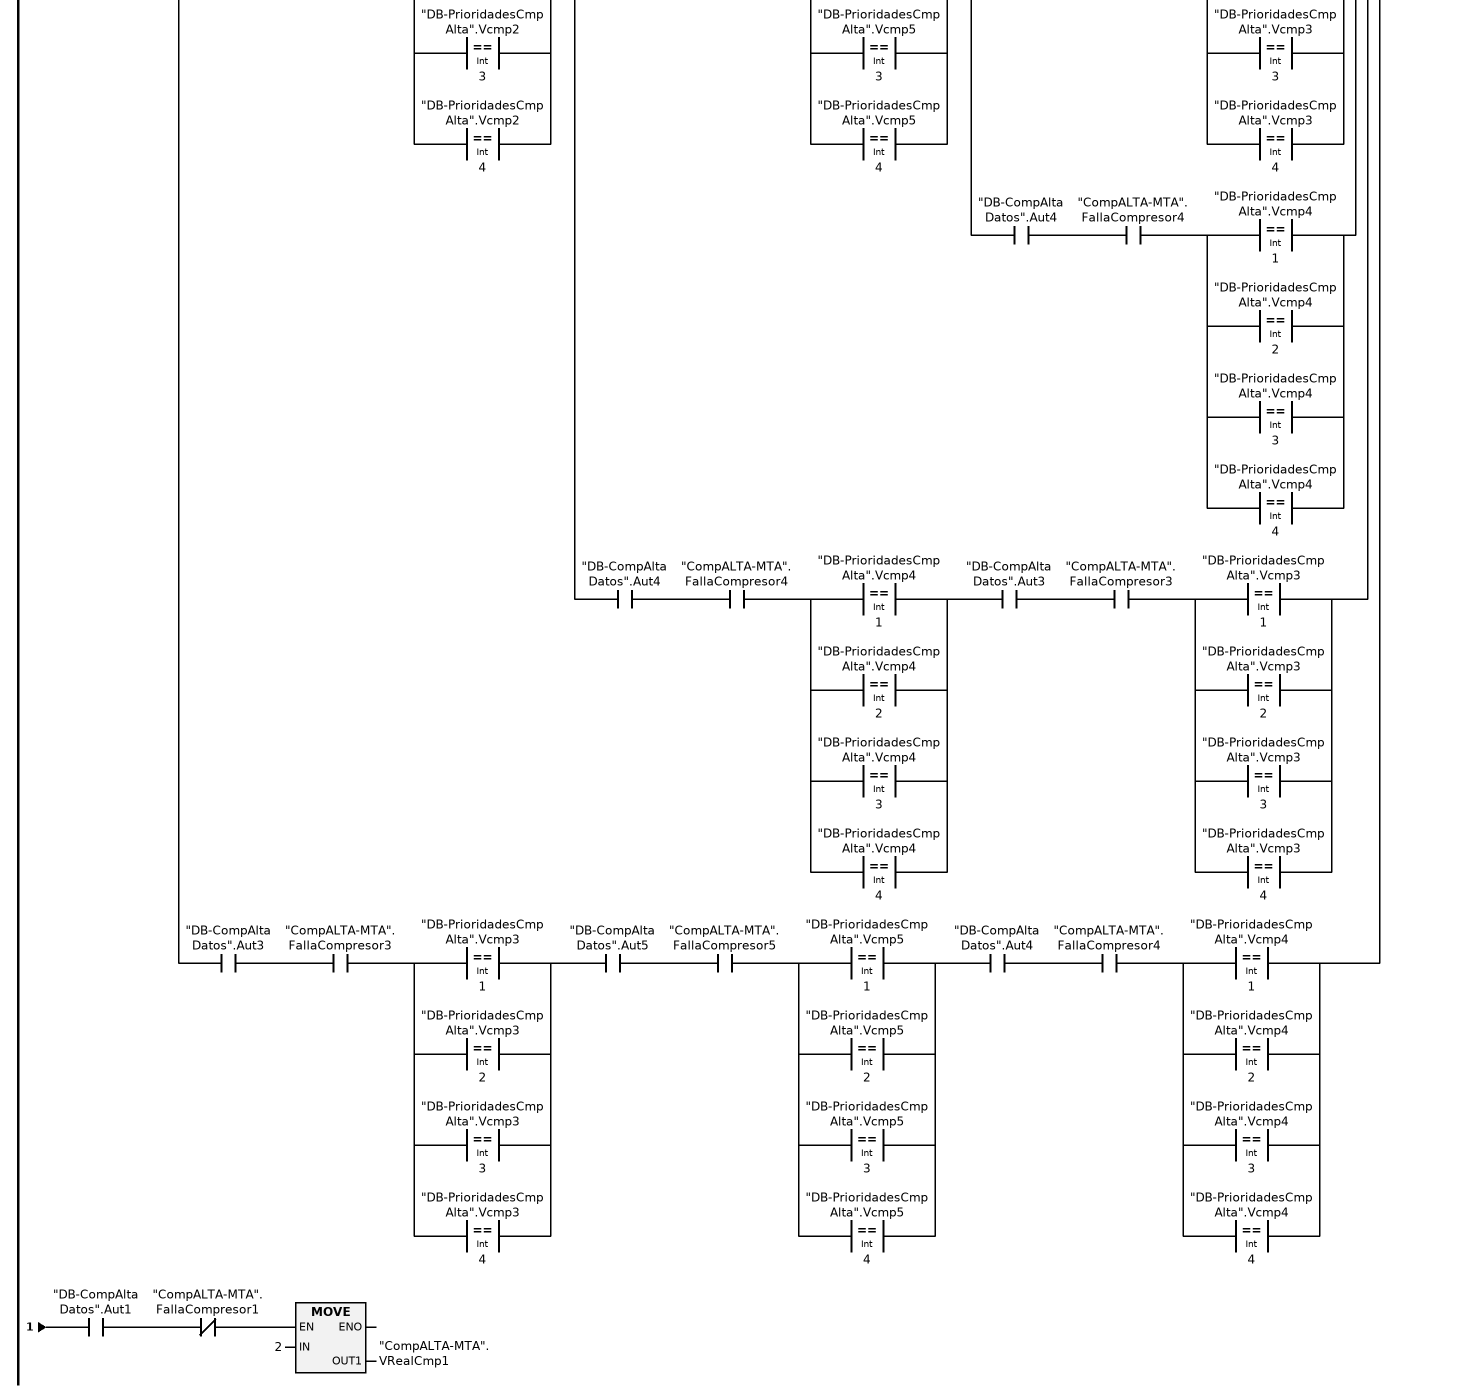
   RUNG wire#powerrail
      { S7_Templates := "SrcType := Int" } EQ_Contact(in1 := "DB-PrioridadesCmpAlta".Vcmp1, in2 := 2)
      wire#w1
      Contact( "DB-CompAltaDatos".Aut1 )
      I_Contact( "CompALTA-MTA".FallaCompresor1 )
      { S7_GenerateENO := "TRUE" } Move(in := 2, out1 => "CompALTA-MTA".VRealCmp1)
   END_RUNG
   RUNG wire#powerrail
      { S7_Templates := "SrcType := Int" } EQ_Contact(in1 := "DB-PrioridadesCmpAlta".Vcmp1, in2 := 3)
      wire#w2
      Contact( "DB-CompAltaDatos".Aut2 )
      Contact( "CompALTA-MTA".FallaCompresor2 )
      wire#w3
      { S7_Templates := "SrcType := Int" } EQ_Contact(in1 := "DB-PrioridadesCmpAlta".Vcmp2, in2 := 2)
   END_RUNG wire#w1
   RUNG wire#w3
      { S7_Templates := "SrcType := Int" } EQ_Contact(in1 := "DB-PrioridadesCmpAlta".Vcmp2, in2 := 1)
   END_RUNG wire#w1
   RUNG wire#w2
      Contact( "DB-CompAltaDatos".Aut3 )
      Contact( "CompALTA-MTA".FallaCompresor3 )
      wire#w4
      { S7_Templates := "SrcType := Int" } EQ_Contact(in1 := "DB-PrioridadesCmpAlta".Vcmp3, in2 := 2)
   END_RUNG wire#w1
   RUNG wire#w4
      { S7_Templates := "SrcType := Int" } EQ_Contact(in1 := "DB-PrioridadesCmpAlta".Vcmp3, in2 := 1)
   END_RUNG wire#w1
   RUNG wire#w2
      Contact( "DB-CompAltaDatos".Aut4 )
      Contact( "CompALTA-MTA".FallaCompresor4 )
      wire#w5
      { S7_Templates := "SrcType := Int" } EQ_Contact(in1 := "DB-PrioridadesCmpAlta".Vcmp4, in2 := 2)
   END_RUNG wire#w1
   RUNG wire#w5
      { S7_Templates := "SrcType := Int" } EQ_Contact(in1 := "DB-PrioridadesCmpAlta".Vcmp4, in2 := 1)
   END_RUNG wire#w1
   RUNG wire#w2
      Contact( "DB-CompAltaDatos".Aut5 )
      Contact( "CompALTA-MTA".FallaCompresor5 )
      wire#w6
      { S7_Templates := "SrcType := Int" } EQ_Contact(in1 := "DB-PrioridadesCmpAlta".Vcmp5, in2 := 2)
   END_RUNG wire#w1
   RUNG wire#w6
      { S7_Templates := "SrcType := Int" } EQ_Contact(in1 := "DB-PrioridadesCmpAlta".Vcmp5, in2 := 1)
   END_RUNG wire#w1
   RUNG wire#powerrail
      { S7_Templates := "SrcType := Int" } EQ_Contact(in1 := "DB-PrioridadesCmpAlta".Vcmp1, in2 := 4)
      wire#w7
      Contact( "DB-CompAltaDatos".Aut2 )
      Contact( "CompALTA-MTA".FallaCompresor2 )
      wire#w8
      { S7_Templates := "SrcType := Int" } EQ_Contact(in1 := "DB-PrioridadesCmpAlta".Vcmp2, in2 := 1)
      wire#w9
      Contact( "DB-CompAltaDatos".Aut5 )
      Contact( "CompALTA-MTA".FallaCompresor5 )
      wire#w10
      { S7_Templates := "SrcType := Int" } EQ_Contact(in1 := "DB-PrioridadesCmpAlta".Vcmp5, in2 := 1)
   END_RUNG wire#w1
   RUNG wire#w8
      { S7_Templates := "SrcType := Int" } EQ_Contact(in1 := "DB-PrioridadesCmpAlta".Vcmp2, in2 := 2)
   END_RUNG wire#w9
   RUNG wire#w8
      { S7_Templates := "SrcType := Int" } EQ_Contact(in1 := "DB-PrioridadesCmpAlta".Vcmp2, in2 := 3)
   END_RUNG wire#w9
   RUNG wire#w10
      { S7_Templates := "SrcType := Int" } EQ_Contact(in1 := "DB-PrioridadesCmpAlta".Vcmp5, in2 := 2)
   END_RUNG wire#w1
   RUNG wire#w10
      { S7_Templates := "SrcType := Int" } EQ_Contact(in1 := "DB-PrioridadesCmpAlta".Vcmp5, in2 := 3)
   END_RUNG wire#w1
   RUNG wire#w9
      Contact( "DB-CompAltaDatos".Aut4 )
      Contact( "CompALTA-MTA".FallaCompresor4 )
      wire#w11
      { S7_Templates := "SrcType := Int" } EQ_Contact(in1 := "DB-PrioridadesCmpAlta".Vcmp4, in2 := 1)
   END_RUNG wire#w1
   RUNG wire#w11
      { S7_Templates := "SrcType := Int" } EQ_Contact(in1 := "DB-PrioridadesCmpAlta".Vcmp4, in2 := 2)
   END_RUNG wire#w1
   RUNG wire#w11
      { S7_Templates := "SrcType := Int" } EQ_Contact(in1 := "DB-PrioridadesCmpAlta".Vcmp4, in2 := 3)
   END_RUNG wire#w1
   RUNG wire#w9
      Contact( "DB-CompAltaDatos".Aut3 )
      Contact( "CompALTA-MTA".FallaCompresor3 )
      wire#w12
      { S7_Templates := "SrcType := Int" } EQ_Contact(in1 := "DB-PrioridadesCmpAlta".Vcmp3, in2 := 1)
   END_RUNG wire#w1
   RUNG wire#w12
      { S7_Templates := "SrcType := Int" } EQ_Contact(in1 := "DB-PrioridadesCmpAlta".Vcmp3, in2 := 2)
   END_RUNG wire#w1
   RUNG wire#w12
      { S7_Templates := "SrcType := Int" } EQ_Contact(in1 := "DB-PrioridadesCmpAlta".Vcmp3, in2 := 3)
   END_RUNG wire#w1
   RUNG wire#w7
      Contact( "DB-CompAltaDatos".Aut3 )
      Contact( "CompALTA-MTA".FallaCompresor3 )
      wire#w13
      { S7_Templates := "SrcType := Int" } EQ_Contact(in1 := "DB-PrioridadesCmpAlta".Vcmp3, in2 := 1)
      wire#w14
      Contact( "DB-CompAltaDatos".Aut5 )
      Contact( "CompALTA-MTA".FallaCompresor5 )
      wire#w15
      { S7_Templates := "SrcType := Int" } EQ_Contact(in1 := "DB-PrioridadesCmpAlta".Vcmp5, in2 := 1)
   END_RUNG wire#w1
   RUNG wire#w13
      { S7_Templates := "SrcType := Int" } EQ_Contact(in1 := "DB-PrioridadesCmpAlta".Vcmp3, in2 := 2)
   END_RUNG wire#w14
   RUNG wire#w13
      { S7_Templates := "SrcType := Int" } EQ_Contact(in1 := "DB-PrioridadesCmpAlta".Vcmp3, in2 := 3)
   END_RUNG wire#w14
   RUNG wire#w15
      { S7_Templates := "SrcType := Int" } EQ_Contact(in1 := "DB-PrioridadesCmpAlta".Vcmp5, in2 := 2)
   END_RUNG wire#w1
   RUNG wire#w15
      { S7_Templates := "SrcType := Int" } EQ_Contact(in1 := "DB-PrioridadesCmpAlta".Vcmp5, in2 := 3)
   END_RUNG wire#w1
   RUNG wire#w14
      Contact( "DB-CompAltaDatos".Aut4 )
      Contact( "CompALTA-MTA".FallaCompresor4 )
      wire#w16
      { S7_Templates := "SrcType := Int" } EQ_Contact(in1 := "DB-PrioridadesCmpAlta".Vcmp4, in2 := 1)
   END_RUNG wire#w1
   RUNG wire#w16
      { S7_Templates := "SrcType := Int" } EQ_Contact(in1 := "DB-PrioridadesCmpAlta".Vcmp4, in2 := 2)
   END_RUNG wire#w1
   RUNG wire#w16
      { S7_Templates := "SrcType := Int" } EQ_Contact(in1 := "DB-PrioridadesCmpAlta".Vcmp4, in2 := 3)
   END_RUNG wire#w1
   RUNG wire#w7
      Contact( "DB-CompAltaDatos".Aut4 )
      Contact( "CompALTA-MTA".FallaCompresor4 )
      wire#w17
      { S7_Templates := "SrcType := Int" } EQ_Contact(in1 := "DB-PrioridadesCmpAlta".Vcmp4, in2 := 1)
      wire#w18
      Contact( "DB-CompAltaDatos".Aut5 )
      Contact( "CompALTA-MTA".FallaCompresor5 )
      wire#w19
      { S7_Templates := "SrcType := Int" } EQ_Contact(in1 := "DB-PrioridadesCmpAlta".Vcmp5, in2 := 1)
   END_RUNG wire#w1
   RUNG wire#w17
      { S7_Templates := "SrcType := Int" } EQ_Contact(in1 := "DB-PrioridadesCmpAlta".Vcmp4, in2 := 2)
   END_RUNG wire#w18
   RUNG wire#w17
      { S7_Templates := "SrcType := Int" } EQ_Contact(in1 := "DB-PrioridadesCmpAlta".Vcmp4, in2 := 3)
   END_RUNG wire#w18
   RUNG wire#w19
      { S7_Templates := "SrcType := Int" } EQ_Contact(in1 := "DB-PrioridadesCmpAlta".Vcmp5, in2 := 2)
   END_RUNG wire#w1
   RUNG wire#w19
      { S7_Templates := "SrcType := Int" } EQ_Contact(in1 := "DB-PrioridadesCmpAlta".Vcmp5, in2 := 3)
   END_RUNG wire#w1
   RUNG wire#powerrail
      { S7_Templates := "SrcType := Int" } EQ_Contact(in1 := "DB-PrioridadesCmpAlta".Vcmp1, in2 := 5)
      wire#w20
      Contact( "DB-CompAltaDatos".Aut2 )
      Contact( "CompALTA-MTA".FallaCompresor2 )
      wire#w21
      { S7_Templates := "SrcType := Int" } EQ_Contact(in1 := "DB-PrioridadesCmpAlta".Vcmp2, in2 := 1)
      wire#w22
      Contact( "DB-CompAltaDatos".Aut5 )
      Contact( "CompALTA-MTA".FallaCompresor5 )
      wire#w23
      { S7_Templates := "SrcType := Int" } EQ_Contact(in1 := "DB-PrioridadesCmpAlta".Vcmp5, in2 := 1)
      wire#w24
      Contact( "DB-CompAltaDatos".Aut3 )
      Contact( "CompALTA-MTA".FallaCompresor3 )
      wire#w25
      { S7_Templates := "SrcType := Int" } EQ_Contact(in1 := "DB-PrioridadesCmpAlta".Vcmp3, in2 := 1)
   END_RUNG wire#w1
   RUNG wire#w21
      { S7_Templates := "SrcType := Int" } EQ_Contact(in1 := "DB-PrioridadesCmpAlta".Vcmp2, in2 := 2)
   END_RUNG wire#w22
   RUNG wire#w21
      { S7_Templates := "SrcType := Int" } EQ_Contact(in1 := "DB-PrioridadesCmpAlta".Vcmp2, in2 := 3)
   END_RUNG wire#w22
   RUNG wire#w21
      { S7_Templates := "SrcType := Int" } EQ_Contact(in1 := "DB-PrioridadesCmpAlta".Vcmp2, in2 := 4)
   END_RUNG wire#w22
   RUNG wire#w23
      { S7_Templates := "SrcType := Int" } EQ_Contact(in1 := "DB-PrioridadesCmpAlta".Vcmp5, in2 := 2)
   END_RUNG wire#w24
   RUNG wire#w23
      { S7_Templates := "SrcType := Int" } EQ_Contact(in1 := "DB-PrioridadesCmpAlta".Vcmp5, in2 := 3)
   END_RUNG wire#w24
   RUNG wire#w23
      { S7_Templates := "SrcType := Int" } EQ_Contact(in1 := "DB-PrioridadesCmpAlta".Vcmp5, in2 := 4)
   END_RUNG wire#w24
   RUNG wire#w25
      { S7_Templates := "SrcType := Int" } EQ_Contact(in1 := "DB-PrioridadesCmpAlta".Vcmp3, in2 := 2)
   END_RUNG wire#w1
   RUNG wire#w25
      { S7_Templates := "SrcType := Int" } EQ_Contact(in1 := "DB-PrioridadesCmpAlta".Vcmp3, in2 := 3)
   END_RUNG wire#w1
   RUNG wire#w25
      { S7_Templates := "SrcType := Int" } EQ_Contact(in1 := "DB-PrioridadesCmpAlta".Vcmp3, in2 := 4)
   END_RUNG wire#w1
   RUNG wire#w24
      Contact( "DB-CompAltaDatos".Aut4 )
      Contact( "CompALTA-MTA".FallaCompresor4 )
      wire#w26
      { S7_Templates := "SrcType := Int" } EQ_Contact(in1 := "DB-PrioridadesCmpAlta".Vcmp4, in2 := 1)
   END_RUNG wire#w1
   RUNG wire#w26
      { S7_Templates := "SrcType := Int" } EQ_Contact(in1 := "DB-PrioridadesCmpAlta".Vcmp4, in2 := 2)
   END_RUNG wire#w1
   RUNG wire#w26
      { S7_Templates := "SrcType := Int" } EQ_Contact(in1 := "DB-PrioridadesCmpAlta".Vcmp4, in2 := 3)
   END_RUNG wire#w1
   RUNG wire#w26
      { S7_Templates := "SrcType := Int" } EQ_Contact(in1 := "DB-PrioridadesCmpAlta".Vcmp4, in2 := 4)
   END_RUNG wire#w1
   RUNG wire#w22
      Contact( "DB-CompAltaDatos".Aut4 )
      Contact( "CompALTA-MTA".FallaCompresor4 )
      wire#w27
      { S7_Templates := "SrcType := Int" } EQ_Contact(in1 := "DB-PrioridadesCmpAlta".Vcmp4, in2 := 1)
      wire#w28
      Contact( "DB-CompAltaDatos".Aut3 )
      Contact( "CompALTA-MTA".FallaCompresor3 )
      wire#w29
      { S7_Templates := "SrcType := Int" } EQ_Contact(in1 := "DB-PrioridadesCmpAlta".Vcmp3, in2 := 1)
   END_RUNG wire#w1
   RUNG wire#w27
      { S7_Templates := "SrcType := Int" } EQ_Contact(in1 := "DB-PrioridadesCmpAlta".Vcmp4, in2 := 2)
   END_RUNG wire#w28
   RUNG wire#w27
      { S7_Templates := "SrcType := Int" } EQ_Contact(in1 := "DB-PrioridadesCmpAlta".Vcmp4, in2 := 3)
   END_RUNG wire#w28
   RUNG wire#w27
      { S7_Templates := "SrcType := Int" } EQ_Contact(in1 := "DB-PrioridadesCmpAlta".Vcmp4, in2 := 4)
   END_RUNG wire#w28
   RUNG wire#w29
      { S7_Templates := "SrcType := Int" } EQ_Contact(in1 := "DB-PrioridadesCmpAlta".Vcmp3, in2 := 2)
   END_RUNG wire#w1
   RUNG wire#w29
      { S7_Templates := "SrcType := Int" } EQ_Contact(in1 := "DB-PrioridadesCmpAlta".Vcmp3, in2 := 3)
   END_RUNG wire#w1
   RUNG wire#w29
      { S7_Templates := "SrcType := Int" } EQ_Contact(in1 := "DB-PrioridadesCmpAlta".Vcmp3, in2 := 4)
   END_RUNG wire#w1
   RUNG wire#w20
      Contact( "DB-CompAltaDatos".Aut3 )
      Contact( "CompALTA-MTA".FallaCompresor3 )
      wire#w30
      { S7_Templates := "SrcType := Int" } EQ_Contact(in1 := "DB-PrioridadesCmpAlta".Vcmp3, in2 := 1)
      wire#w31
      Contact( "DB-CompAltaDatos".Aut5 )
      Contact( "CompALTA-MTA".FallaCompresor5 )
      wire#w32
      { S7_Templates := "SrcType := Int" } EQ_Contact(in1 := "DB-PrioridadesCmpAlta".Vcmp5, in2 := 1)
      wire#w33
      Contact( "DB-CompAltaDatos".Aut4 )
      Contact( "CompALTA-MTA".FallaCompresor4 )
      wire#w34
      { S7_Templates := "SrcType := Int" } EQ_Contact(in1 := "DB-PrioridadesCmpAlta".Vcmp4, in2 := 1)
   END_RUNG wire#w1
   RUNG wire#w30
      { S7_Templates := "SrcType := Int" } EQ_Contact(in1 := "DB-PrioridadesCmpAlta".Vcmp3, in2 := 2)
   END_RUNG wire#w31
   RUNG wire#w30
      { S7_Templates := "SrcType := Int" } EQ_Contact(in1 := "DB-PrioridadesCmpAlta".Vcmp3, in2 := 3)
   END_RUNG wire#w31
   RUNG wire#w30
      { S7_Templates := "SrcType := Int" } EQ_Contact(in1 := "DB-PrioridadesCmpAlta".Vcmp3, in2 := 4)
   END_RUNG wire#w31
   RUNG wire#w32
      { S7_Templates := "SrcType := Int" } EQ_Contact(in1 := "DB-PrioridadesCmpAlta".Vcmp5, in2 := 2)
   END_RUNG wire#w33
   RUNG wire#w32
      { S7_Templates := "SrcType := Int" } EQ_Contact(in1 := "DB-PrioridadesCmpAlta".Vcmp5, in2 := 3)
   END_RUNG wire#w33
   RUNG wire#w32
      { S7_Templates := "SrcType := Int" } EQ_Contact(in1 := "DB-PrioridadesCmpAlta".Vcmp5, in2 := 4)
   END_RUNG wire#w33
   RUNG wire#w34
      { S7_Templates := "SrcType := Int" } EQ_Contact(in1 := "DB-PrioridadesCmpAlta".Vcmp4, in2 := 2)
   END_RUNG wire#w1
   RUNG wire#w34
      { S7_Templates := "SrcType := Int" } EQ_Contact(in1 := "DB-PrioridadesCmpAlta".Vcmp4, in2 := 3)
   END_RUNG wire#w1
   RUNG wire#w34
      { S7_Templates := "SrcType := Int" } EQ_Contact(in1 := "DB-PrioridadesCmpAlta".Vcmp4, in2 := 4)
   END_RUNG wire#w1
   // the same network as SCL:
   IF (("DB-PrioridadesCmpAlta".Vcmp1 = 2) OR (("DB-PrioridadesCmpAlta".Vcmp1 = 3) AND (("DB-CompAltaDatos".Aut2 AND "CompALTA-MTA".FallaCompresor2 AND (("DB-PrioridadesCmpAlta".Vcmp2 = 2) OR ("DB-PrioridadesCmpAlta".Vcmp2 = 1))) OR ("DB-CompAltaDatos".Aut3 AND "CompALTA-MTA".FallaCompresor3 AND (("DB-PrioridadesCmpAlta".Vcmp3 = 2) OR ("DB-PrioridadesCmpAlta".Vcmp3 = 1))) OR ("DB-CompAltaDatos".Aut4 AND "CompALTA-MTA".FallaCompresor4 AND (("DB-PrioridadesCmpAlta".Vcmp4 = 2) OR ("DB-PrioridadesCmpAlta".Vcmp4 = 1))) OR ("DB-CompAltaDatos".Aut5 AND "CompALTA-MTA".FallaCompresor5 AND (("DB-PrioridadesCmpAlta".Vcmp5 = 2) OR ("DB-PrioridadesCmpAlta".Vcmp5 = 1))))) OR (("DB-PrioridadesCmpAlta".Vcmp1 = 4) AND (("DB-CompAltaDatos".Aut2 AND "CompALTA-MTA".FallaCompresor2 AND (("DB-PrioridadesCmpAlta".Vcmp2 = 1) OR ("DB-PrioridadesCmpAlta".Vcmp2 = 2) OR ("DB-PrioridadesCmpAlta".Vcmp2 = 3)) AND (("DB-CompAltaDatos".Aut5 AND "CompALTA-MTA".FallaCompresor5 AND (("DB-PrioridadesCmpAlta".Vcmp5 = 1) OR ("DB-PrioridadesCmpAlta".Vcmp5 = 2) OR ("DB-PrioridadesCmpAlta".Vcmp5 = 3))) OR ("DB-CompAltaDatos".Aut4 AND "CompALTA-MTA".FallaCompresor4 AND (("DB-PrioridadesCmpAlta".Vcmp4 = 1) OR ("DB-PrioridadesCmpAlta".Vcmp4 = 2) OR ("DB-PrioridadesCmpAlta".Vcmp4 = 3))) OR ("DB-CompAltaDatos".Aut3 AND "CompALTA-MTA".FallaCompresor3 AND (("DB-PrioridadesCmpAlta".Vcmp3 = 1) OR ("DB-PrioridadesCmpAlta".Vcmp3 = 2) OR ("DB-PrioridadesCmpAlta".Vcmp3 = 3))))) OR ("DB-CompAltaDatos".Aut3 AND "CompALTA-MTA".FallaCompresor3 AND (("DB-PrioridadesCmpAlta".Vcmp3 = 1) OR ("DB-PrioridadesCmpAlta".Vcmp3 = 2) OR ("DB-PrioridadesCmpAlta".Vcmp3 = 3)) AND (("DB-CompAltaDatos".Aut5 AND "CompALTA-MTA".FallaCompresor5 AND (("DB-PrioridadesCmpAlta".Vcmp5 = 1) OR ("DB-PrioridadesCmpAlta".Vcmp5 = 2) OR ("DB-PrioridadesCmpAlta".Vcmp5 = 3))) OR ("DB-CompAltaDatos".Aut4 AND "CompALTA-MTA".FallaCompresor4 AND (("DB-PrioridadesCmpAlta".Vcmp4 = 1) OR ("DB-PrioridadesCmpAlta".Vcmp4 = 2) OR ("DB-PrioridadesCmpAlta".Vcmp4 = 3))))) OR ("DB-CompAltaDatos".Aut4 AND "CompALTA-MTA".FallaCompresor4 AND (("DB-PrioridadesCmpAlta".Vcmp4 = 1) OR ("DB-PrioridadesCmpAlta".Vcmp4 = 2) OR ("DB-PrioridadesCmpAlta".Vcmp4 = 3)) AND "DB-CompAltaDatos".Aut5 AND "CompALTA-MTA".FallaCompresor5 AND (("DB-PrioridadesCmpAlta".Vcmp5 = 1) OR ("DB-PrioridadesCmpAlta".Vcmp5 = 2) OR ("DB-PrioridadesCmpAlta".Vcmp5 = 3))))) OR (("DB-PrioridadesCmpAlta".Vcmp1 = 5) AND (("DB-CompAltaDatos".Aut2 AND "CompALTA-MTA".FallaCompresor2 AND (("DB-PrioridadesCmpAlta".Vcmp2 = 1) OR ("DB-PrioridadesCmpAlta".Vcmp2 = 2) OR ("DB-PrioridadesCmpAlta".Vcmp2 = 3) OR ("DB-PrioridadesCmpAlta".Vcmp2 = 4)) AND (("DB-CompAltaDatos".Aut5 AND "CompALTA-MTA".FallaCompresor5 AND (("DB-PrioridadesCmpAlta".Vcmp5 = 1) OR ("DB-PrioridadesCmpAlta".Vcmp5 = 2) OR ("DB-PrioridadesCmpAlta".Vcmp5 = 3) OR ("DB-PrioridadesCmpAlta".Vcmp5 = 4)) AND (("DB-CompAltaDatos".Aut3 AND "CompALTA-MTA".FallaCompresor3 AND (("DB-PrioridadesCmpAlta".Vcmp3 = 1) OR ("DB-PrioridadesCmpAlta".Vcmp3 = 2) OR ("DB-PrioridadesCmpAlta".Vcmp3 = 3) OR ("DB-PrioridadesCmpAlta".Vcmp3 = 4))) OR ("DB-CompAltaDatos".Aut4 AND "CompALTA-MTA".FallaCompresor4 AND (("DB-PrioridadesCmpAlta".Vcmp4 = 1) OR ("DB-PrioridadesCmpAlta".Vcmp4 = 2) OR ("DB-PrioridadesCmpAlta".Vcmp4 = 3) OR ("DB-PrioridadesCmpAlta".Vcmp4 = 4))))) OR ("DB-CompAltaDatos".Aut4 AND "CompALTA-MTA".FallaCompresor4 AND (("DB-PrioridadesCmpAlta".Vcmp4 = 1) OR ("DB-PrioridadesCmpAlta".Vcmp4 = 2) OR ("DB-PrioridadesCmpAlta".Vcmp4 = 3) OR ("DB-PrioridadesCmpAlta".Vcmp4 = 4)) AND "DB-CompAltaDatos".Aut3 AND "CompALTA-MTA".FallaCompresor3 AND (("DB-PrioridadesCmpAlta".Vcmp3 = 1) OR ("DB-PrioridadesCmpAlta".Vcmp3 = 2) OR ("DB-PrioridadesCmpAlta".Vcmp3 = 3) OR ("DB-PrioridadesCmpAlta".Vcmp3 = 4))))) OR ("DB-CompAltaDatos".Aut3 AND "CompALTA-MTA".FallaCompresor3 AND (("DB-PrioridadesCmpAlta".Vcmp3 = 1) OR ("DB-PrioridadesCmpAlta".Vcmp3 = 2) OR ("DB-PrioridadesCmpAlta".Vcmp3 = 3) OR ("DB-PrioridadesCmpAlta".Vcmp3 = 4)) AND "DB-CompAltaDatos".Aut5 AND "CompALTA-MTA".FallaCompresor5 AND (("DB-PrioridadesCmpAlta".Vcmp5 = 1) OR ("DB-PrioridadesCmpAlta".Vcmp5 = 2) OR ("DB-PrioridadesCmpAlta".Vcmp5 = 3) OR ("DB-PrioridadesCmpAlta".Vcmp5 = 4)) AND "DB-CompAltaDatos".Aut4 AND "CompALTA-MTA".FallaCompresor4 AND (("DB-PrioridadesCmpAlta".Vcmp4 = 1) OR ("DB-PrioridadesCmpAlta".Vcmp4 = 2) OR ("DB-PrioridadesCmpAlta".Vcmp4 = 3) OR ("DB-PrioridadesCmpAlta".Vcmp4 = 4)))))) AND "DB-CompAltaDatos".Aut1 AND NOT "CompALTA-MTA".FallaCompresor1 THEN
       "CompALTA-MTA".VRealCmp1 := 2;
   END_IF;
END_REGION

REGION Network 5
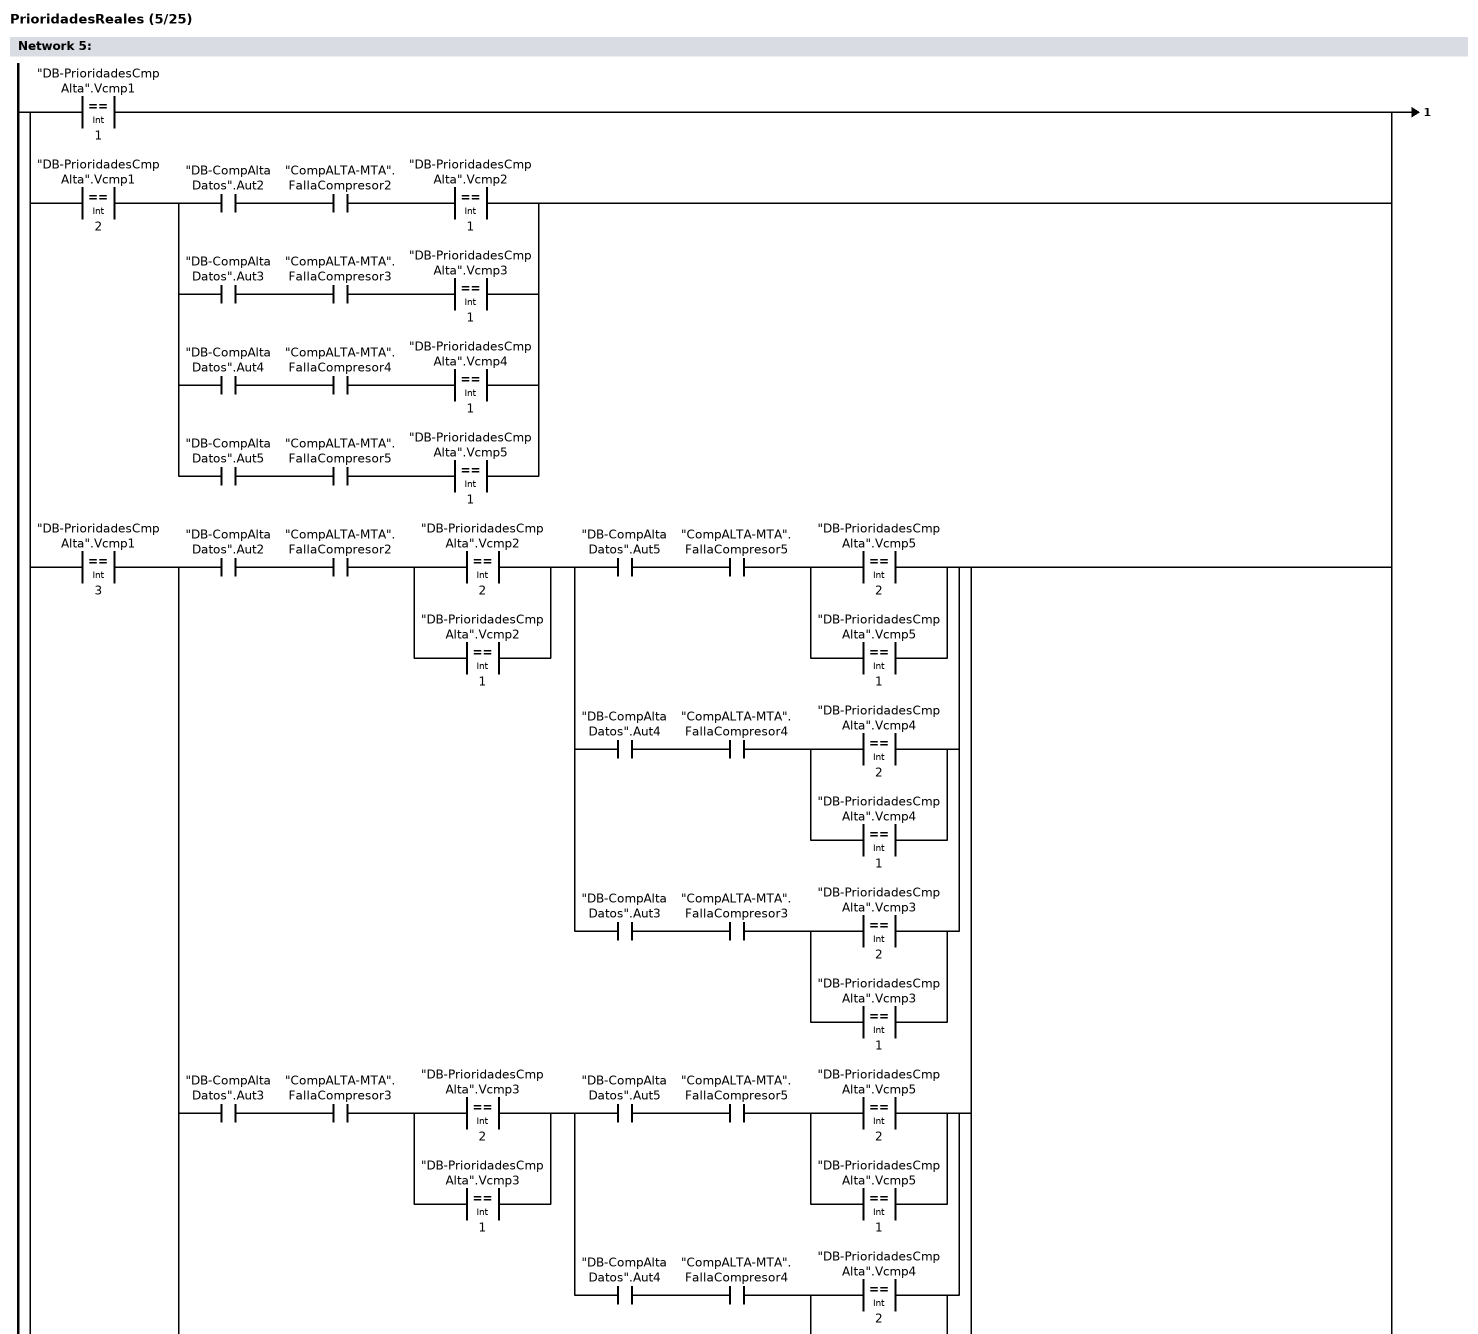
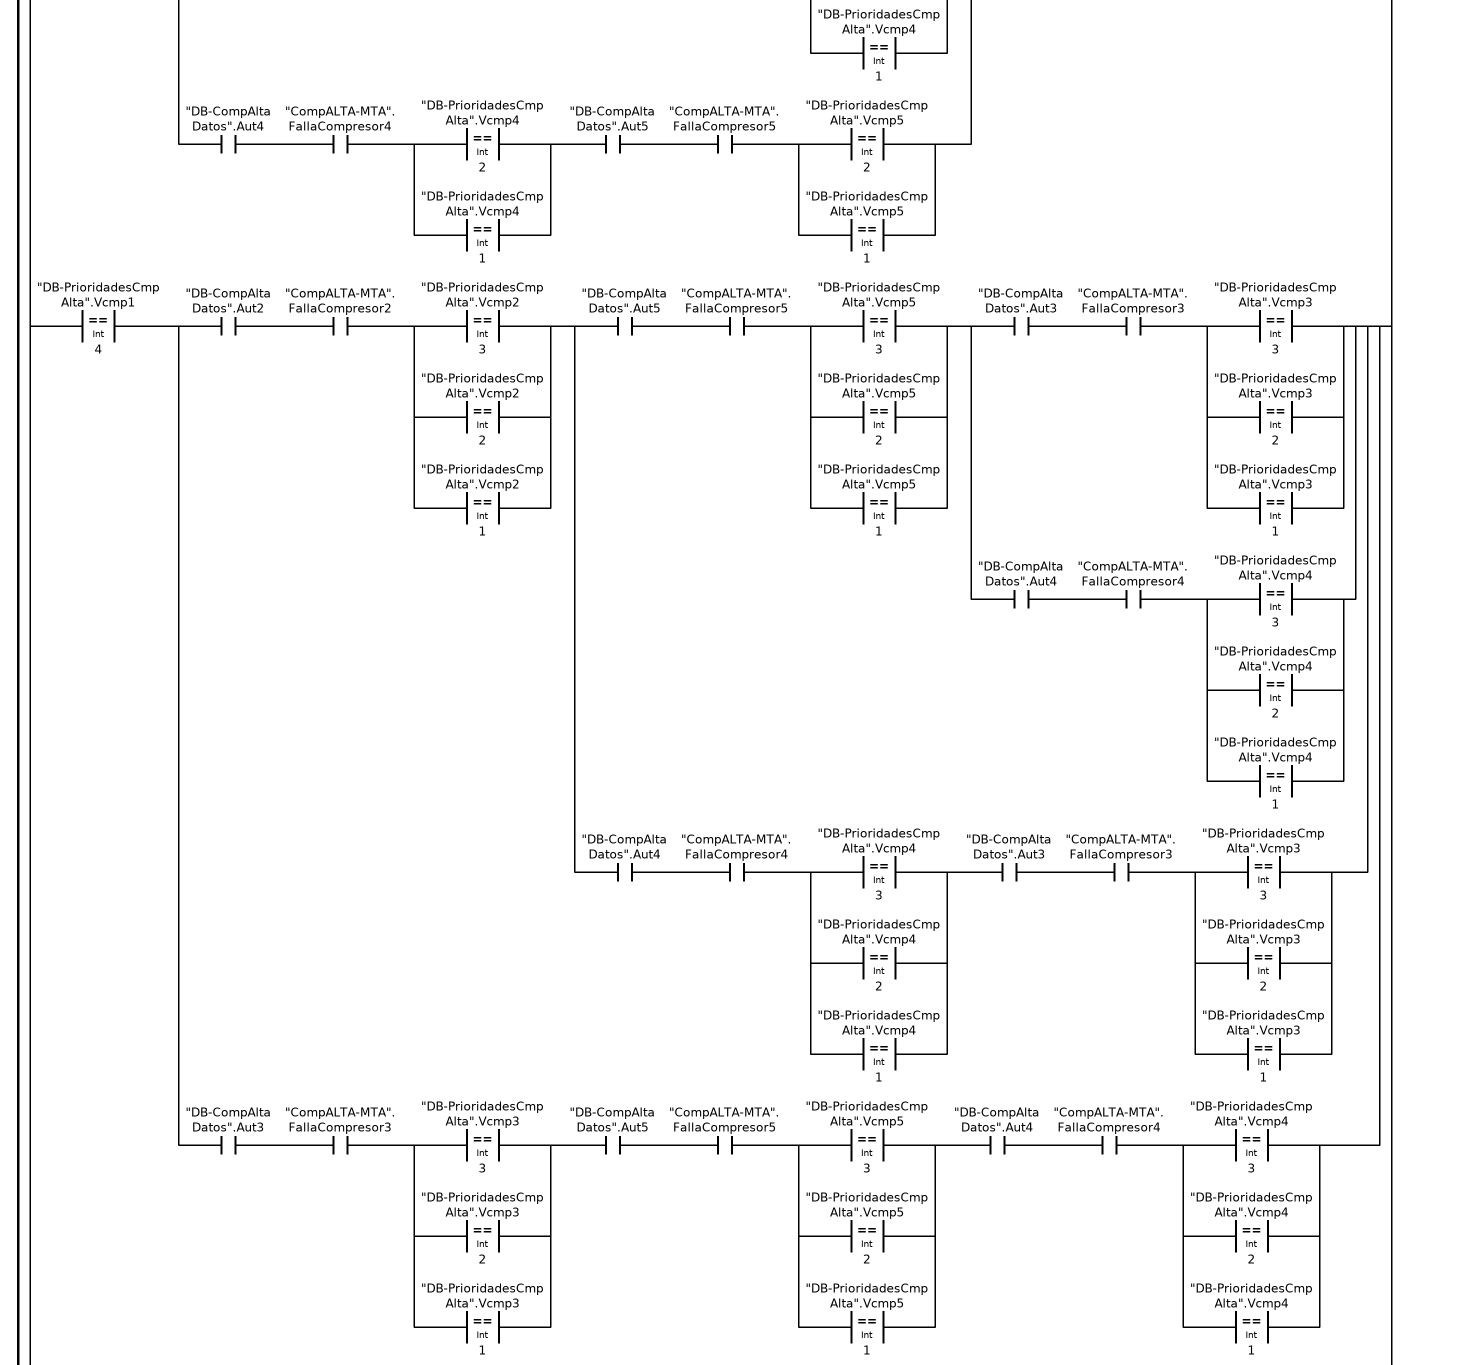
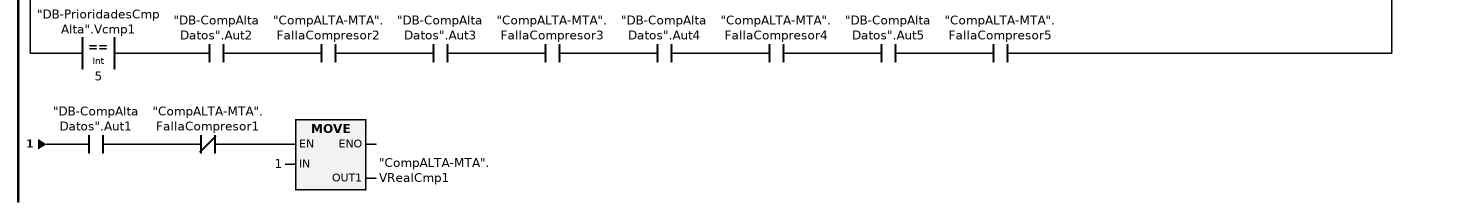
   RUNG wire#powerrail
      { S7_Templates := "SrcType := Int" } EQ_Contact(in1 := "DB-PrioridadesCmpAlta".Vcmp1, in2 := 1)
      wire#w1
      Contact( "DB-CompAltaDatos".Aut1 )
      I_Contact( "CompALTA-MTA".FallaCompresor1 )
      { S7_GenerateENO := "TRUE" } Move(in := 1, out1 => "CompALTA-MTA".VRealCmp1)
   END_RUNG
   RUNG wire#powerrail
      { S7_Templates := "SrcType := Int" } EQ_Contact(in1 := "DB-PrioridadesCmpAlta".Vcmp1, in2 := 2)
      wire#w2
      Contact( "DB-CompAltaDatos".Aut2 )
      Contact( "CompALTA-MTA".FallaCompresor2 )
      { S7_Templates := "SrcType := Int" } EQ_Contact(in1 := "DB-PrioridadesCmpAlta".Vcmp2, in2 := 1)
   END_RUNG wire#w1
   RUNG wire#w2
      Contact( "DB-CompAltaDatos".Aut3 )
      Contact( "CompALTA-MTA".FallaCompresor3 )
      { S7_Templates := "SrcType := Int" } EQ_Contact(in1 := "DB-PrioridadesCmpAlta".Vcmp3, in2 := 1)
   END_RUNG wire#w1
   RUNG wire#w2
      Contact( "DB-CompAltaDatos".Aut4 )
      Contact( "CompALTA-MTA".FallaCompresor4 )
      { S7_Templates := "SrcType := Int" } EQ_Contact(in1 := "DB-PrioridadesCmpAlta".Vcmp4, in2 := 1)
   END_RUNG wire#w1
   RUNG wire#w2
      Contact( "DB-CompAltaDatos".Aut5 )
      Contact( "CompALTA-MTA".FallaCompresor5 )
      { S7_Templates := "SrcType := Int" } EQ_Contact(in1 := "DB-PrioridadesCmpAlta".Vcmp5, in2 := 1)
   END_RUNG wire#w1
   RUNG wire#powerrail
      { S7_Templates := "SrcType := Int" } EQ_Contact(in1 := "DB-PrioridadesCmpAlta".Vcmp1, in2 := 3)
      wire#w3
      Contact( "DB-CompAltaDatos".Aut2 )
      Contact( "CompALTA-MTA".FallaCompresor2 )
      wire#w4
      { S7_Templates := "SrcType := Int" } EQ_Contact(in1 := "DB-PrioridadesCmpAlta".Vcmp2, in2 := 2)
      wire#w5
      Contact( "DB-CompAltaDatos".Aut5 )
      Contact( "CompALTA-MTA".FallaCompresor5 )
      wire#w6
      { S7_Templates := "SrcType := Int" } EQ_Contact(in1 := "DB-PrioridadesCmpAlta".Vcmp5, in2 := 2)
   END_RUNG wire#w1
   RUNG wire#w4
      { S7_Templates := "SrcType := Int" } EQ_Contact(in1 := "DB-PrioridadesCmpAlta".Vcmp2, in2 := 1)
   END_RUNG wire#w5
   RUNG wire#w6
      { S7_Templates := "SrcType := Int" } EQ_Contact(in1 := "DB-PrioridadesCmpAlta".Vcmp5, in2 := 1)
   END_RUNG wire#w1
   RUNG wire#w5
      Contact( "DB-CompAltaDatos".Aut4 )
      Contact( "CompALTA-MTA".FallaCompresor4 )
      wire#w7
      { S7_Templates := "SrcType := Int" } EQ_Contact(in1 := "DB-PrioridadesCmpAlta".Vcmp4, in2 := 2)
   END_RUNG wire#w1
   RUNG wire#w7
      { S7_Templates := "SrcType := Int" } EQ_Contact(in1 := "DB-PrioridadesCmpAlta".Vcmp4, in2 := 1)
   END_RUNG wire#w1
   RUNG wire#w5
      Contact( "DB-CompAltaDatos".Aut3 )
      Contact( "CompALTA-MTA".FallaCompresor3 )
      wire#w8
      { S7_Templates := "SrcType := Int" } EQ_Contact(in1 := "DB-PrioridadesCmpAlta".Vcmp3, in2 := 2)
   END_RUNG wire#w1
   RUNG wire#w8
      { S7_Templates := "SrcType := Int" } EQ_Contact(in1 := "DB-PrioridadesCmpAlta".Vcmp3, in2 := 1)
   END_RUNG wire#w1
   RUNG wire#w3
      Contact( "DB-CompAltaDatos".Aut3 )
      Contact( "CompALTA-MTA".FallaCompresor3 )
      wire#w9
      { S7_Templates := "SrcType := Int" } EQ_Contact(in1 := "DB-PrioridadesCmpAlta".Vcmp3, in2 := 2)
      wire#w10
      Contact( "DB-CompAltaDatos".Aut5 )
      Contact( "CompALTA-MTA".FallaCompresor5 )
      wire#w11
      { S7_Templates := "SrcType := Int" } EQ_Contact(in1 := "DB-PrioridadesCmpAlta".Vcmp5, in2 := 2)
   END_RUNG wire#w1
   RUNG wire#w9
      { S7_Templates := "SrcType := Int" } EQ_Contact(in1 := "DB-PrioridadesCmpAlta".Vcmp3, in2 := 1)
   END_RUNG wire#w10
   RUNG wire#w11
      { S7_Templates := "SrcType := Int" } EQ_Contact(in1 := "DB-PrioridadesCmpAlta".Vcmp5, in2 := 1)
   END_RUNG wire#w1
   RUNG wire#w10
      Contact( "DB-CompAltaDatos".Aut4 )
      Contact( "CompALTA-MTA".FallaCompresor4 )
      wire#w12
      { S7_Templates := "SrcType := Int" } EQ_Contact(in1 := "DB-PrioridadesCmpAlta".Vcmp4, in2 := 2)
   END_RUNG wire#w1
   RUNG wire#w12
      { S7_Templates := "SrcType := Int" } EQ_Contact(in1 := "DB-PrioridadesCmpAlta".Vcmp4, in2 := 1)
   END_RUNG wire#w1
   RUNG wire#w3
      Contact( "DB-CompAltaDatos".Aut4 )
      Contact( "CompALTA-MTA".FallaCompresor4 )
      wire#w13
      { S7_Templates := "SrcType := Int" } EQ_Contact(in1 := "DB-PrioridadesCmpAlta".Vcmp4, in2 := 2)
      wire#w14
      Contact( "DB-CompAltaDatos".Aut5 )
      Contact( "CompALTA-MTA".FallaCompresor5 )
      wire#w15
      { S7_Templates := "SrcType := Int" } EQ_Contact(in1 := "DB-PrioridadesCmpAlta".Vcmp5, in2 := 2)
   END_RUNG wire#w1
   RUNG wire#w13
      { S7_Templates := "SrcType := Int" } EQ_Contact(in1 := "DB-PrioridadesCmpAlta".Vcmp4, in2 := 1)
   END_RUNG wire#w14
   RUNG wire#w15
      { S7_Templates := "SrcType := Int" } EQ_Contact(in1 := "DB-PrioridadesCmpAlta".Vcmp5, in2 := 1)
   END_RUNG wire#w1
   RUNG wire#powerrail
      { S7_Templates := "SrcType := Int" } EQ_Contact(in1 := "DB-PrioridadesCmpAlta".Vcmp1, in2 := 4)
      wire#w16
      Contact( "DB-CompAltaDatos".Aut2 )
      Contact( "CompALTA-MTA".FallaCompresor2 )
      wire#w17
      { S7_Templates := "SrcType := Int" } EQ_Contact(in1 := "DB-PrioridadesCmpAlta".Vcmp2, in2 := 3)
      wire#w18
      Contact( "DB-CompAltaDatos".Aut5 )
      Contact( "CompALTA-MTA".FallaCompresor5 )
      wire#w19
      { S7_Templates := "SrcType := Int" } EQ_Contact(in1 := "DB-PrioridadesCmpAlta".Vcmp5, in2 := 3)
      wire#w20
      Contact( "DB-CompAltaDatos".Aut3 )
      Contact( "CompALTA-MTA".FallaCompresor3 )
      wire#w21
      { S7_Templates := "SrcType := Int" } EQ_Contact(in1 := "DB-PrioridadesCmpAlta".Vcmp3, in2 := 3)
   END_RUNG wire#w1
   RUNG wire#w17
      { S7_Templates := "SrcType := Int" } EQ_Contact(in1 := "DB-PrioridadesCmpAlta".Vcmp2, in2 := 2)
   END_RUNG wire#w18
   RUNG wire#w17
      { S7_Templates := "SrcType := Int" } EQ_Contact(in1 := "DB-PrioridadesCmpAlta".Vcmp2, in2 := 1)
   END_RUNG wire#w18
   RUNG wire#w19
      { S7_Templates := "SrcType := Int" } EQ_Contact(in1 := "DB-PrioridadesCmpAlta".Vcmp5, in2 := 2)
   END_RUNG wire#w20
   RUNG wire#w19
      { S7_Templates := "SrcType := Int" } EQ_Contact(in1 := "DB-PrioridadesCmpAlta".Vcmp5, in2 := 1)
   END_RUNG wire#w20
   RUNG wire#w21
      { S7_Templates := "SrcType := Int" } EQ_Contact(in1 := "DB-PrioridadesCmpAlta".Vcmp3, in2 := 2)
   END_RUNG wire#w1
   RUNG wire#w21
      { S7_Templates := "SrcType := Int" } EQ_Contact(in1 := "DB-PrioridadesCmpAlta".Vcmp3, in2 := 1)
   END_RUNG wire#w1
   RUNG wire#w20
      Contact( "DB-CompAltaDatos".Aut4 )
      Contact( "CompALTA-MTA".FallaCompresor4 )
      wire#w22
      { S7_Templates := "SrcType := Int" } EQ_Contact(in1 := "DB-PrioridadesCmpAlta".Vcmp4, in2 := 3)
   END_RUNG wire#w1
   RUNG wire#w22